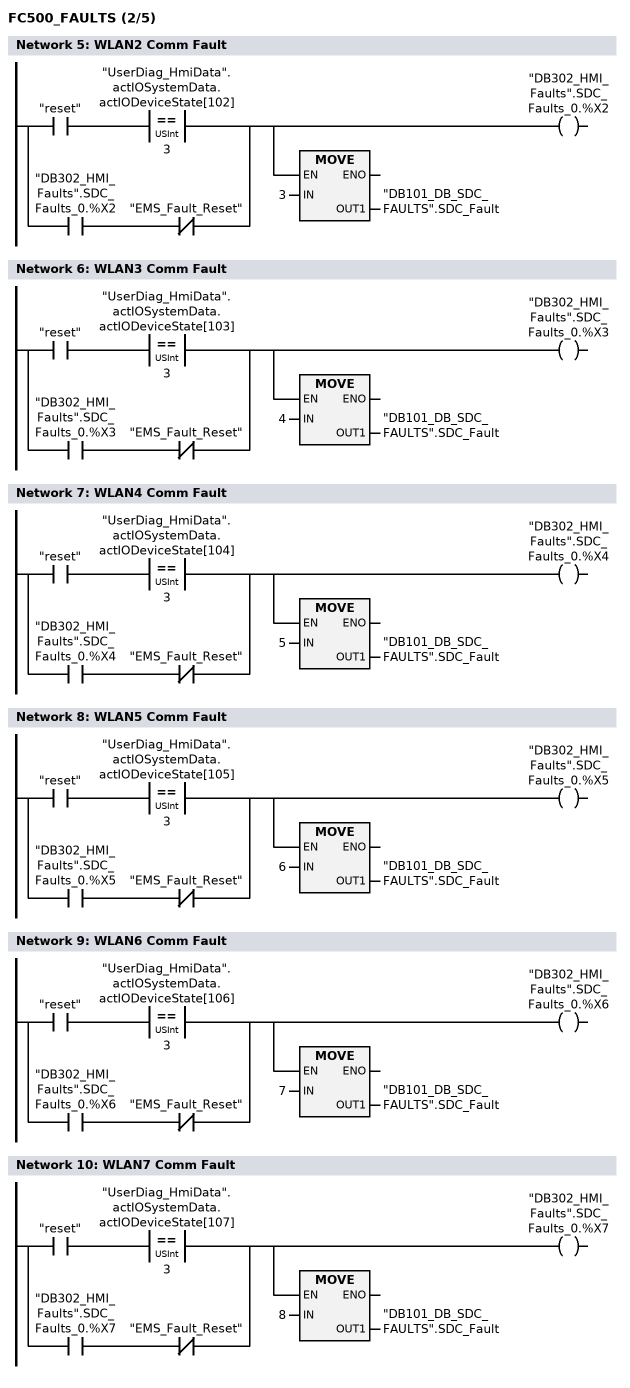
   RUNG wire#powerrail
      Contact( "reset" )
      { S7_Templates := "SrcType := USInt" } EQ_Contact(in1 := "UserDiag_HmiData".actIOSystemData.actIODeviceState[102], in2 := 3)
      wire#w1
      Coil( "DB302_HMI_Faults".SDC_Faults_0.%X2 )
   END_RUNG
   RUNG wire#powerrail
      Contact( "DB302_HMI_Faults".SDC_Faults_0.%X2 )
      I_Contact( "EMS_Fault_Reset" )
   END_RUNG wire#w1
   RUNG wire#w1
      Move(in := 3, out1 => "DB101_DB_SDC_FAULTS".SDC_Fault)
   END_RUNG
   // the same network as SCL:
   "DB302_HMI_Faults".SDC_Faults_0.%X2 := ("reset" AND ("UserDiag_HmiData".actIOSystemData.actIODeviceState[102] = 3)) OR ("DB302_HMI_Faults".SDC_Faults_0.%X2 AND NOT "EMS_Fault_Reset");
   IF "DB302_HMI_Faults".SDC_Faults_0.%X2 THEN "DB101_DB_SDC_FAULTS".SDC_Fault := 3; END_IF;
END_REGION

REGION Network 6: WLAN3 Comm Fault
   RUNG wire#powerrail
      Contact( "reset" )
      { S7_Templates := "SrcType := USInt" } EQ_Contact(in1 := "UserDiag_HmiData".actIOSystemData.actIODeviceState[103], in2 := 3)
      wire#w1
      Coil( "DB302_HMI_Faults".SDC_Faults_0.%X3 )
   END_RUNG
   RUNG wire#powerrail
      Contact( "DB302_HMI_Faults".SDC_Faults_0.%X3 )
      I_Contact( "EMS_Fault_Reset" )
   END_RUNG wire#w1
   RUNG wire#w1
      Move(in := 4, out1 => "DB101_DB_SDC_FAULTS".SDC_Fault)
   END_RUNG
   // the same network as SCL:
   "DB302_HMI_Faults".SDC_Faults_0.%X3 := ("reset" AND ("UserDiag_HmiData".actIOSystemData.actIODeviceState[103] = 3)) OR ("DB302_HMI_Faults".SDC_Faults_0.%X3 AND NOT "EMS_Fault_Reset");
   IF "DB302_HMI_Faults".SDC_Faults_0.%X3 THEN "DB101_DB_SDC_FAULTS".SDC_Fault := 4; END_IF;
END_REGION

REGION Network 7: WLAN4 Comm Fault
   RUNG wire#powerrail
      Contact( "reset" )
      { S7_Templates := "SrcType := USInt" } EQ_Contact(in1 := "UserDiag_HmiData".actIOSystemData.actIODeviceState[104], in2 := 3)
      wire#w1
      Coil( "DB302_HMI_Faults".SDC_Faults_0.%X4 )
   END_RUNG
   RUNG wire#powerrail
      Contact( "DB302_HMI_Faults".SDC_Faults_0.%X4 )
      I_Contact( "EMS_Fault_Reset" )
   END_RUNG wire#w1
   RUNG wire#w1
      Move(in := 5, out1 => "DB101_DB_SDC_FAULTS".SDC_Fault)
   END_RUNG
   // the same network as SCL:
   "DB302_HMI_Faults".SDC_Faults_0.%X4 := ("reset" AND ("UserDiag_HmiData".actIOSystemData.actIODeviceState[104] = 3)) OR ("DB302_HMI_Faults".SDC_Faults_0.%X4 AND NOT "EMS_Fault_Reset");
   IF "DB302_HMI_Faults".SDC_Faults_0.%X4 THEN "DB101_DB_SDC_FAULTS".SDC_Fault := 5; END_IF;
END_REGION

REGION Network 8: WLAN5 Comm Fault
   RUNG wire#powerrail
      Contact( "reset" )
      { S7_Templates := "SrcType := USInt" } EQ_Contact(in1 := "UserDiag_HmiData".actIOSystemData.actIODeviceState[105], in2 := 3)
      wire#w1
      Coil( "DB302_HMI_Faults".SDC_Faults_0.%X5 )
   END_RUNG
   RUNG wire#powerrail
      Contact( "DB302_HMI_Faults".SDC_Faults_0.%X5 )
      I_Contact( "EMS_Fault_Reset" )
   END_RUNG wire#w1
   RUNG wire#w1
      Move(in := 6, out1 => "DB101_DB_SDC_FAULTS".SDC_Fault)
   END_RUNG
   // the same network as SCL:
   "DB302_HMI_Faults".SDC_Faults_0.%X5 := ("reset" AND ("UserDiag_HmiData".actIOSystemData.actIODeviceState[105] = 3)) OR ("DB302_HMI_Faults".SDC_Faults_0.%X5 AND NOT "EMS_Fault_Reset");
   IF "DB302_HMI_Faults".SDC_Faults_0.%X5 THEN "DB101_DB_SDC_FAULTS".SDC_Fault := 6; END_IF;
END_REGION

REGION Network 9: WLAN6 Comm Fault
   RUNG wire#powerrail
      Contact( "reset" )
      { S7_Templates := "SrcType := USInt" } EQ_Contact(in1 := "UserDiag_HmiData".actIOSystemData.actIODeviceState[106], in2 := 3)
      wire#w1
      Coil( "DB302_HMI_Faults".SDC_Faults_0.%X6 )
   END_RUNG
   RUNG wire#powerrail
      Contact( "DB302_HMI_Faults".SDC_Faults_0.%X6 )
      I_Contact( "EMS_Fault_Reset" )
   END_RUNG wire#w1
   RUNG wire#w1
      Move(in := 7, out1 => "DB101_DB_SDC_FAULTS".SDC_Fault)
   END_RUNG
   // the same network as SCL:
   "DB302_HMI_Faults".SDC_Faults_0.%X6 := ("reset" AND ("UserDiag_HmiData".actIOSystemData.actIODeviceState[106] = 3)) OR ("DB302_HMI_Faults".SDC_Faults_0.%X6 AND NOT "EMS_Fault_Reset");
   IF "DB302_HMI_Faults".SDC_Faults_0.%X6 THEN "DB101_DB_SDC_FAULTS".SDC_Fault := 7; END_IF;
END_REGION

REGION Network 10: WLAN7 Comm Fault
   RUNG wire#powerrail
      Contact( "reset" )
      { S7_Templates := "SrcType := USInt" } EQ_Contact(in1 := "UserDiag_HmiData".actIOSystemData.actIODeviceState[107], in2 := 3)
      wire#w1
      Coil( "DB302_HMI_Faults".SDC_Faults_0.%X7 )
   END_RUNG
   RUNG wire#powerrail
      Contact( "DB302_HMI_Faults".SDC_Faults_0.%X7 )
      I_Contact( "EMS_Fault_Reset" )
   END_RUNG wire#w1
   RUNG wire#w1
      Move(in := 8, out1 => "DB101_DB_SDC_FAULTS".SDC_Fault)
   END_RUNG
   // the same network as SCL:
   "DB302_HMI_Faults".SDC_Faults_0.%X7 := ("reset" AND ("UserDiag_HmiData".actIOSystemData.actIODeviceState[107] = 3)) OR ("DB302_HMI_Faults".SDC_Faults_0.%X7 AND NOT "EMS_Fault_Reset");
   IF "DB302_HMI_Faults".SDC_Faults_0.%X7 THEN "DB101_DB_SDC_FAULTS".SDC_Fault := 8; END_IF;
END_REGION

REGION Network 11: WLAN8 Comm Fault
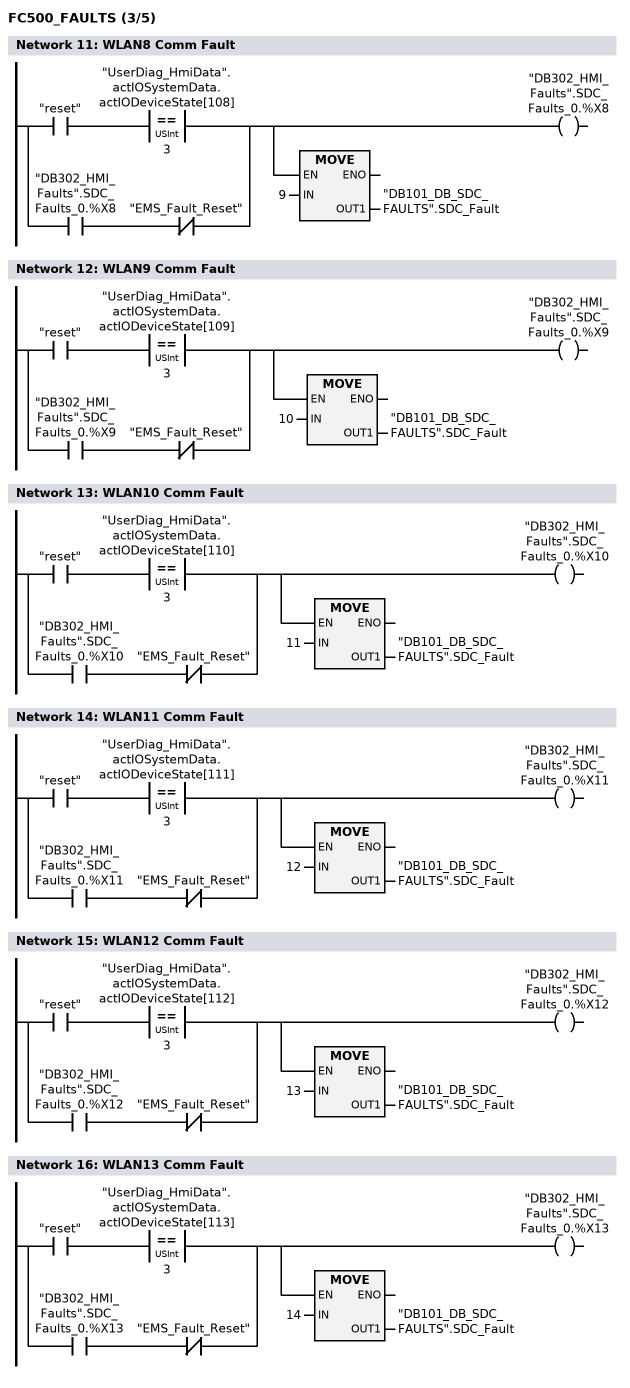
   RUNG wire#powerrail
      Contact( "reset" )
      { S7_Templates := "SrcType := USInt" } EQ_Contact(in1 := "UserDiag_HmiData".actIOSystemData.actIODeviceState[108], in2 := 3)
      wire#w1
      Coil( "DB302_HMI_Faults".SDC_Faults_0.%X8 )
   END_RUNG
   RUNG wire#powerrail
      Contact( "DB302_HMI_Faults".SDC_Faults_0.%X8 )
      I_Contact( "EMS_Fault_Reset" )
   END_RUNG wire#w1
   RUNG wire#w1
      Move(in := 9, out1 => "DB101_DB_SDC_FAULTS".SDC_Fault)
   END_RUNG
   // the same network as SCL:
   "DB302_HMI_Faults".SDC_Faults_0.%X8 := ("reset" AND ("UserDiag_HmiData".actIOSystemData.actIODeviceState[108] = 3)) OR ("DB302_HMI_Faults".SDC_Faults_0.%X8 AND NOT "EMS_Fault_Reset");
   IF "DB302_HMI_Faults".SDC_Faults_0.%X8 THEN "DB101_DB_SDC_FAULTS".SDC_Fault := 9; END_IF;
END_REGION

REGION Network 12: WLAN9 Comm Fault
   RUNG wire#powerrail
      Contact( "reset" )
      { S7_Templates := "SrcType := USInt" } EQ_Contact(in1 := "UserDiag_HmiData".actIOSystemData.actIODeviceState[109], in2 := 3)
      wire#w1
      Coil( "DB302_HMI_Faults".SDC_Faults_0.%X9 )
   END_RUNG
   RUNG wire#powerrail
      Contact( "DB302_HMI_Faults".SDC_Faults_0.%X9 )
      I_Contact( "EMS_Fault_Reset" )
   END_RUNG wire#w1
   RUNG wire#w1
      Move(in := 10, out1 => "DB101_DB_SDC_FAULTS".SDC_Fault)
   END_RUNG
   // the same network as SCL:
   "DB302_HMI_Faults".SDC_Faults_0.%X9 := ("reset" AND ("UserDiag_HmiData".actIOSystemData.actIODeviceState[109] = 3)) OR ("DB302_HMI_Faults".SDC_Faults_0.%X9 AND NOT "EMS_Fault_Reset");
   IF "DB302_HMI_Faults".SDC_Faults_0.%X9 THEN "DB101_DB_SDC_FAULTS".SDC_Fault := 10; END_IF;
END_REGION

REGION Network 13: WLAN10 Comm Fault
   RUNG wire#powerrail
      Contact( "reset" )
      { S7_Templates := "SrcType := USInt" } EQ_Contact(in1 := "UserDiag_HmiData".actIOSystemData.actIODeviceState[110], in2 := 3)
      wire#w1
      Coil( "DB302_HMI_Faults".SDC_Faults_0.%X10 )
   END_RUNG
   RUNG wire#powerrail
      Contact( "DB302_HMI_Faults".SDC_Faults_0.%X10 )
      I_Contact( "EMS_Fault_Reset" )
   END_RUNG wire#w1
   RUNG wire#w1
      Move(in := 11, out1 => "DB101_DB_SDC_FAULTS".SDC_Fault)
   END_RUNG
   // the same network as SCL:
   "DB302_HMI_Faults".SDC_Faults_0.%X10 := ("reset" AND ("UserDiag_HmiData".actIOSystemData.actIODeviceState[110] = 3)) OR ("DB302_HMI_Faults".SDC_Faults_0.%X10 AND NOT "EMS_Fault_Reset");
   IF "DB302_HMI_Faults".SDC_Faults_0.%X10 THEN "DB101_DB_SDC_FAULTS".SDC_Fault := 11; END_IF;
END_REGION

REGION Network 14: WLAN11 Comm Fault
   RUNG wire#powerrail
      Contact( "reset" )
      { S7_Templates := "SrcType := USInt" } EQ_Contact(in1 := "UserDiag_HmiData".actIOSystemData.actIODeviceState[111], in2 := 3)
      wire#w1
      Coil( "DB302_HMI_Faults".SDC_Faults_0.%X11 )
   END_RUNG
   RUNG wire#powerrail
      Contact( "DB302_HMI_Faults".SDC_Faults_0.%X11 )
      I_Contact( "EMS_Fault_Reset" )
   END_RUNG wire#w1
   RUNG wire#w1
      Move(in := 12, out1 => "DB101_DB_SDC_FAULTS".SDC_Fault)
   END_RUNG
   // the same network as SCL:
   "DB302_HMI_Faults".SDC_Faults_0.%X11 := ("reset" AND ("UserDiag_HmiData".actIOSystemData.actIODeviceState[111] = 3)) OR ("DB302_HMI_Faults".SDC_Faults_0.%X11 AND NOT "EMS_Fault_Reset");
   IF "DB302_HMI_Faults".SDC_Faults_0.%X11 THEN "DB101_DB_SDC_FAULTS".SDC_Fault := 12; END_IF;
END_REGION

REGION Network 15: WLAN12 Comm Fault
   RUNG wire#powerrail
      Contact( "reset" )
      { S7_Templates := "SrcType := USInt" } EQ_Contact(in1 := "UserDiag_HmiData".actIOSystemData.actIODeviceState[112], in2 := 3)
      wire#w1
      Coil( "DB302_HMI_Faults".SDC_Faults_0.%X12 )
   END_RUNG
   RUNG wire#powerrail
      Contact( "DB302_HMI_Faults".SDC_Faults_0.%X12 )
      I_Contact( "EMS_Fault_Reset" )
   END_RUNG wire#w1
   RUNG wire#w1
      Move(in := 13, out1 => "DB101_DB_SDC_FAULTS".SDC_Fault)
   END_RUNG
   // the same network as SCL:
   "DB302_HMI_Faults".SDC_Faults_0.%X12 := ("reset" AND ("UserDiag_HmiData".actIOSystemData.actIODeviceState[112] = 3)) OR ("DB302_HMI_Faults".SDC_Faults_0.%X12 AND NOT "EMS_Fault_Reset");
   IF "DB302_HMI_Faults".SDC_Faults_0.%X12 THEN "DB101_DB_SDC_FAULTS".SDC_Fault := 13; END_IF;
END_REGION

REGION Network 16: WLAN13 Comm Fault
   RUNG wire#powerrail
      Contact( "reset" )
      { S7_Templates := "SrcType := USInt" } EQ_Contact(in1 := "UserDiag_HmiData".actIOSystemData.actIODeviceState[113], in2 := 3)
      wire#w1
      Coil( "DB302_HMI_Faults".SDC_Faults_0.%X13 )
   END_RUNG
   RUNG wire#powerrail
      Contact( "DB302_HMI_Faults".SDC_Faults_0.%X13 )
      I_Contact( "EMS_Fault_Reset" )
   END_RUNG wire#w1
   RUNG wire#w1
      Move(in := 14, out1 => "DB101_DB_SDC_FAULTS".SDC_Fault)
   END_RUNG
   // the same network as SCL:
   "DB302_HMI_Faults".SDC_Faults_0.%X13 := ("reset" AND ("UserDiag_HmiData".actIOSystemData.actIODeviceState[113] = 3)) OR ("DB302_HMI_Faults".SDC_Faults_0.%X13 AND NOT "EMS_Fault_Reset");
   IF "DB302_HMI_Faults".SDC_Faults_0.%X13 THEN "DB101_DB_SDC_FAULTS".SDC_Fault := 14; END_IF;
END_REGION

REGION Network 17: WLAN14 Comm Fault
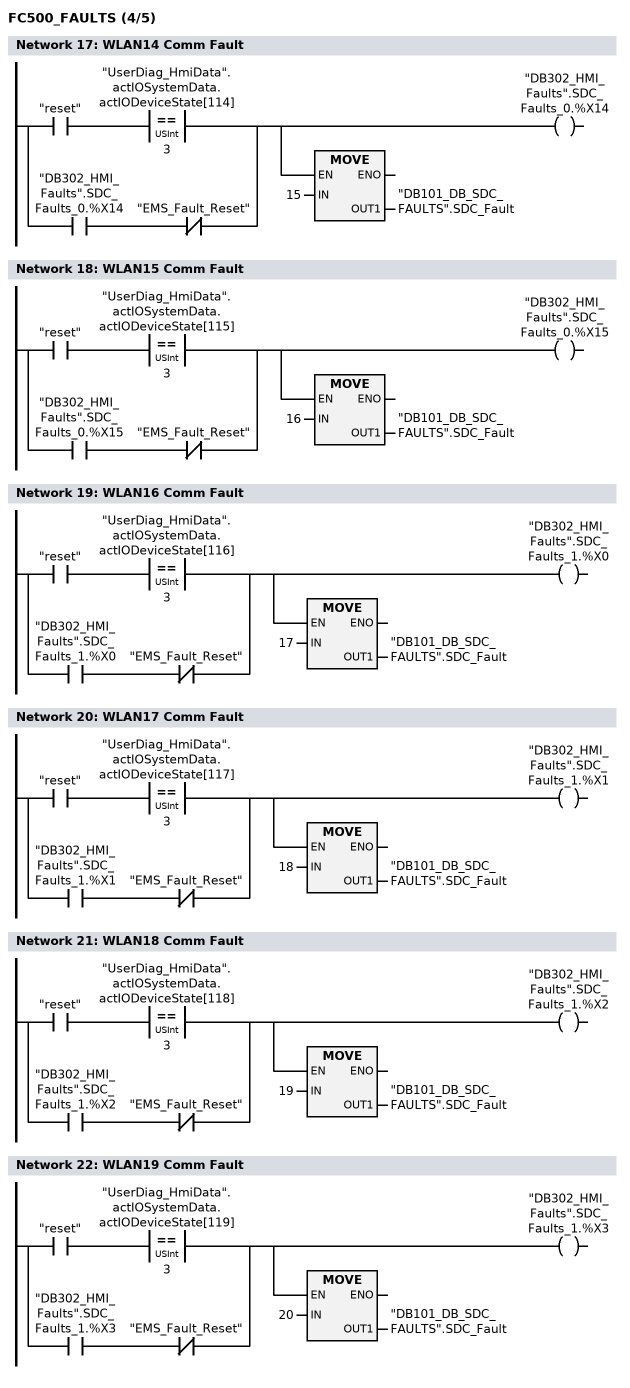
   RUNG wire#powerrail
      Contact( "reset" )
      { S7_Templates := "SrcType := USInt" } EQ_Contact(in1 := "UserDiag_HmiData".actIOSystemData.actIODeviceState[114], in2 := 3)
      wire#w1
      Coil( "DB302_HMI_Faults".SDC_Faults_0.%X14 )
   END_RUNG
   RUNG wire#powerrail
      Contact( "DB302_HMI_Faults".SDC_Faults_0.%X14 )
      I_Contact( "EMS_Fault_Reset" )
   END_RUNG wire#w1
   RUNG wire#w1
      Move(in := 15, out1 => "DB101_DB_SDC_FAULTS".SDC_Fault)
   END_RUNG
   // the same network as SCL:
   "DB302_HMI_Faults".SDC_Faults_0.%X14 := ("reset" AND ("UserDiag_HmiData".actIOSystemData.actIODeviceState[114] = 3)) OR ("DB302_HMI_Faults".SDC_Faults_0.%X14 AND NOT "EMS_Fault_Reset");
   IF "DB302_HMI_Faults".SDC_Faults_0.%X14 THEN "DB101_DB_SDC_FAULTS".SDC_Fault := 15; END_IF;
END_REGION

REGION Network 18: WLAN15 Comm Fault
   RUNG wire#powerrail
      Contact( "reset" )
      { S7_Templates := "SrcType := USInt" } EQ_Contact(in1 := "UserDiag_HmiData".actIOSystemData.actIODeviceState[115], in2 := 3)
      wire#w1
      Coil( "DB302_HMI_Faults".SDC_Faults_0.%X15 )
   END_RUNG
   RUNG wire#powerrail
      Contact( "DB302_HMI_Faults".SDC_Faults_0.%X15 )
      I_Contact( "EMS_Fault_Reset" )
   END_RUNG wire#w1
   RUNG wire#w1
      Move(in := 16, out1 => "DB101_DB_SDC_FAULTS".SDC_Fault)
   END_RUNG
   // the same network as SCL:
   "DB302_HMI_Faults".SDC_Faults_0.%X15 := ("reset" AND ("UserDiag_HmiData".actIOSystemData.actIODeviceState[115] = 3)) OR ("DB302_HMI_Faults".SDC_Faults_0.%X15 AND NOT "EMS_Fault_Reset");
   IF "DB302_HMI_Faults".SDC_Faults_0.%X15 THEN "DB101_DB_SDC_FAULTS".SDC_Fault := 16; END_IF;
END_REGION

REGION Network 19: WLAN16 Comm Fault
   RUNG wire#powerrail
      Contact( "reset" )
      { S7_Templates := "SrcType := USInt" } EQ_Contact(in1 := "UserDiag_HmiData".actIOSystemData.actIODeviceState[116], in2 := 3)
      wire#w1
      Coil( "DB302_HMI_Faults".SDC_Faults_1.%X0 )
   END_RUNG
   RUNG wire#powerrail
      Contact( "DB302_HMI_Faults".SDC_Faults_1.%X0 )
      I_Contact( "EMS_Fault_Reset" )
   END_RUNG wire#w1
   RUNG wire#w1
      Move(in := 17, out1 => "DB101_DB_SDC_FAULTS".SDC_Fault)
   END_RUNG
   // the same network as SCL:
   "DB302_HMI_Faults".SDC_Faults_1.%X0 := ("reset" AND ("UserDiag_HmiData".actIOSystemData.actIODeviceState[116] = 3)) OR ("DB302_HMI_Faults".SDC_Faults_1.%X0 AND NOT "EMS_Fault_Reset");
   IF "DB302_HMI_Faults".SDC_Faults_1.%X0 THEN "DB101_DB_SDC_FAULTS".SDC_Fault := 17; END_IF;
END_REGION

REGION Network 20: WLAN17 Comm Fault
   RUNG wire#powerrail
      Contact( "reset" )
      { S7_Templates := "SrcType := USInt" } EQ_Contact(in1 := "UserDiag_HmiData".actIOSystemData.actIODeviceState[117], in2 := 3)
      wire#w1
      Coil( "DB302_HMI_Faults".SDC_Faults_1.%X1 )
   END_RUNG
   RUNG wire#powerrail
      Contact( "DB302_HMI_Faults".SDC_Faults_1.%X1 )
      I_Contact( "EMS_Fault_Reset" )
   END_RUNG wire#w1
   RUNG wire#w1
      Move(in := 18, out1 => "DB101_DB_SDC_FAULTS".SDC_Fault)
   END_RUNG
   // the same network as SCL:
   "DB302_HMI_Faults".SDC_Faults_1.%X1 := ("reset" AND ("UserDiag_HmiData".actIOSystemData.actIODeviceState[117] = 3)) OR ("DB302_HMI_Faults".SDC_Faults_1.%X1 AND NOT "EMS_Fault_Reset");
   IF "DB302_HMI_Faults".SDC_Faults_1.%X1 THEN "DB101_DB_SDC_FAULTS".SDC_Fault := 18; END_IF;
END_REGION

REGION Network 21: WLAN18 Comm Fault
   RUNG wire#powerrail
      Contact( "reset" )
      { S7_Templates := "SrcType := USInt" } EQ_Contact(in1 := "UserDiag_HmiData".actIOSystemData.actIODeviceState[118], in2 := 3)
      wire#w1
      Coil( "DB302_HMI_Faults".SDC_Faults_1.%X2 )
   END_RUNG
   RUNG wire#powerrail
      Contact( "DB302_HMI_Faults".SDC_Faults_1.%X2 )
      I_Contact( "EMS_Fault_Reset" )
   END_RUNG wire#w1
   RUNG wire#w1
      Move(in := 19, out1 => "DB101_DB_SDC_FAULTS".SDC_Fault)
   END_RUNG
   // the same network as SCL:
   "DB302_HMI_Faults".SDC_Faults_1.%X2 := ("reset" AND ("UserDiag_HmiData".actIOSystemData.actIODeviceState[118] = 3)) OR ("DB302_HMI_Faults".SDC_Faults_1.%X2 AND NOT "EMS_Fault_Reset");
   IF "DB302_HMI_Faults".SDC_Faults_1.%X2 THEN "DB101_DB_SDC_FAULTS".SDC_Fault := 19; END_IF;
END_REGION

REGION Network 22: WLAN19 Comm Fault
   RUNG wire#powerrail
      Contact( "reset" )
      { S7_Templates := "SrcType := USInt" } EQ_Contact(in1 := "UserDiag_HmiData".actIOSystemData.actIODeviceState[119], in2 := 3)
      wire#w1
      Coil( "DB302_HMI_Faults".SDC_Faults_1.%X3 )
   END_RUNG
   RUNG wire#powerrail
      Contact( "DB302_HMI_Faults".SDC_Faults_1.%X3 )
      I_Contact( "EMS_Fault_Reset" )
   END_RUNG wire#w1
   RUNG wire#w1
      Move(in := 20, out1 => "DB101_DB_SDC_FAULTS".SDC_Fault)
   END_RUNG
   // the same network as SCL:
   "DB302_HMI_Faults".SDC_Faults_1.%X3 := ("reset" AND ("UserDiag_HmiData".actIOSystemData.actIODeviceState[119] = 3)) OR ("DB302_HMI_Faults".SDC_Faults_1.%X3 AND NOT "EMS_Fault_Reset");
   IF "DB302_HMI_Faults".SDC_Faults_1.%X3 THEN "DB101_DB_SDC_FAULTS".SDC_Fault := 20; END_IF;
END_REGION

REGION Network 23: Duplicate Carrier Fault
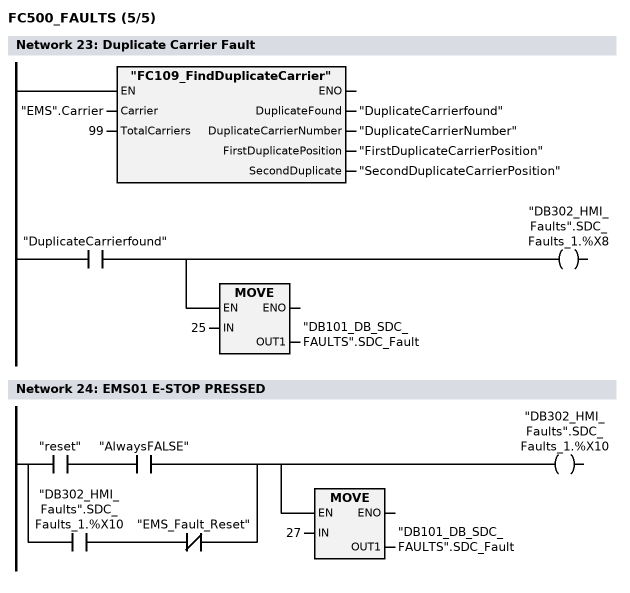
   RUNG wire#powerrail
      "FC109_FindDuplicateCarrier"(Carrier := "EMS".Carrier, TotalCarriers := 99, DuplicateFound => "DuplicateCarrierfound", DuplicateCarrierNumber => "DuplicateCarrierNumber", FirstDuplicatePosition => "FirstDuplicateCarrierPosition", SecondDuplicate => "SecondDuplicateCarrierPosition")
   END_RUNG
   RUNG wire#powerrail
      Contact( "DuplicateCarrierfound" )
      wire#w1
      Coil( "DB302_HMI_Faults".SDC_Faults_1.%X8 )
   END_RUNG
   RUNG wire#w1
      Move(in := 25, out1 => "DB101_DB_SDC_FAULTS".SDC_Fault)
   END_RUNG
   // the same network as SCL:
   "FC109_FindDuplicateCarrier"(Carrier := "EMS".Carrier,
                           TotalCarriers := 99,
                           DuplicateFound => "DuplicateCarrierfound",
                           DuplicateCarrierNumber => "DuplicateCarrierNumber",
                           FirstDuplicatePosition => "FirstDuplicateCarrierPosition",
                           SecondDuplicate => "SecondDuplicateCarrierPosition");
   "DB302_HMI_Faults".SDC_Faults_1.%X8 := "DuplicateCarrierfound";
   IF "DuplicateCarrierfound" THEN "DB101_DB_SDC_FAULTS".SDC_Fault := 25; END_IF;
END_REGION

REGION Network 24: EMS01 E-STOP PRESSED
   RUNG wire#powerrail
      Contact( "reset" )
      Contact( "AlwaysFALSE" )
      wire#w1
      Coil( "DB302_HMI_Faults".SDC_Faults_1.%X10 )
   END_RUNG
   RUNG wire#powerrail
      Contact( "DB302_HMI_Faults".SDC_Faults_1.%X10 )
      I_Contact( "EMS_Fault_Reset" )
   END_RUNG wire#w1
   RUNG wire#w1
      Move(in := 27, out1 => "DB101_DB_SDC_FAULTS".SDC_Fault)
   END_RUNG
   // the same network as SCL:
   "DB302_HMI_Faults".SDC_Faults_1.%X10 := ("reset" AND "AlwaysFALSE") OR ("DB302_HMI_Faults".SDC_Faults_1.%X10 AND NOT "EMS_Fault_Reset");
   IF "DB302_HMI_Faults".SDC_Faults_1.%X10 THEN "DB101_DB_SDC_FAULTS".SDC_Fault := 27; END_IF;
END_REGION
END_FUNCTION

FUNCTION "FC501_FAULTS  C1-C10" : Void   // FC501, LAD
{ S7_Optimized_Access := 'TRUE' }
VERSION : 0.1
BEGIN

REGION Network 1: CARRIER 1 FAULTS
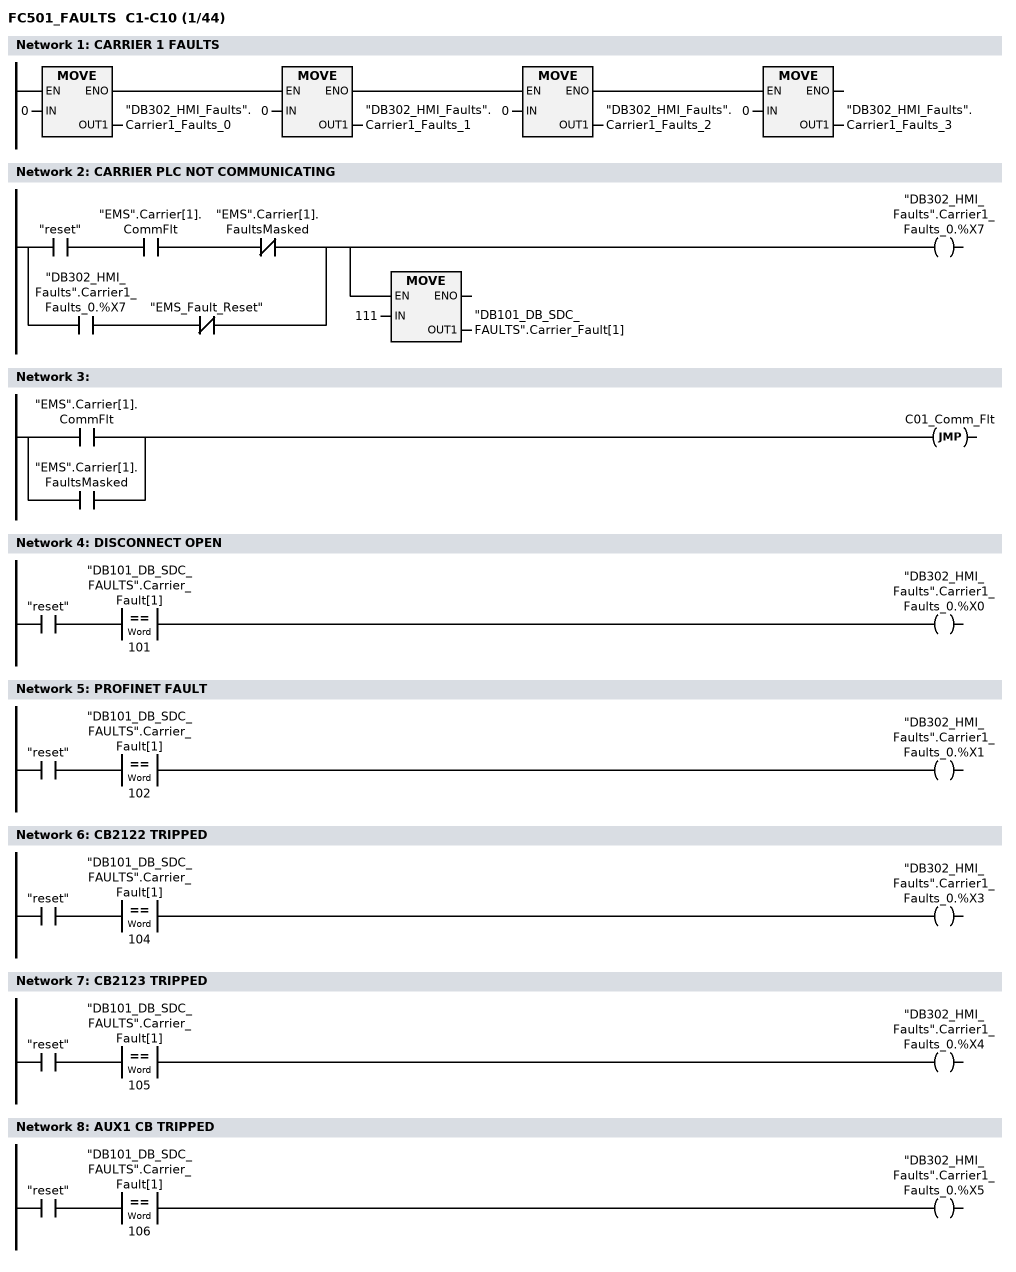
   RUNG wire#powerrail
      Move(in := 0, out1 => "DB302_HMI_Faults".Carrier1_Faults_0)
      Move(in := 0, out1 => "DB302_HMI_Faults".Carrier1_Faults_1)
      Move(in := 0, out1 => "DB302_HMI_Faults".Carrier1_Faults_2)
      Move(in := 0, out1 => "DB302_HMI_Faults".Carrier1_Faults_3)
   END_RUNG
   // the same network as SCL:
   "DB302_HMI_Faults".Carrier1_Faults_0 := 0;
   "DB302_HMI_Faults".Carrier1_Faults_1 := 0;
   "DB302_HMI_Faults".Carrier1_Faults_2 := 0;
   "DB302_HMI_Faults".Carrier1_Faults_3 := 0;
END_REGION

REGION Network 2: CARRIER PLC NOT COMMUNICATING
   RUNG wire#powerrail
      Contact( "reset" )
      Contact( "EMS".Carrier[1].CommFlt )
      I_Contact( "EMS".Carrier[1].FaultsMasked )
      wire#w1
      Coil( "DB302_HMI_Faults".Carrier1_Faults_0.%X7 )
   END_RUNG
   RUNG wire#powerrail
      Contact( "DB302_HMI_Faults".Carrier1_Faults_0.%X7 )
      I_Contact( "EMS_Fault_Reset" )
   END_RUNG wire#w1
   RUNG wire#w1
      Move(in := 111, out1 => "DB101_DB_SDC_FAULTS".Carrier_Fault[1])
   END_RUNG
   // the same network as SCL:
   "DB302_HMI_Faults".Carrier1_Faults_0.%X7 := ("reset" AND "EMS".Carrier[1].CommFlt AND NOT "EMS".Carrier[1].FaultsMasked) OR ("DB302_HMI_Faults".Carrier1_Faults_0.%X7 AND NOT "EMS_Fault_Reset");
   IF "DB302_HMI_Faults".Carrier1_Faults_0.%X7 THEN "DB101_DB_SDC_FAULTS".Carrier_Fault[1] := 111; END_IF;
END_REGION

REGION Network 3
   RUNG wire#powerrail
      Contact( "EMS".Carrier[1].CommFlt )
      wire#w1
      JumpCoil( C01_Comm_Flt )
   END_RUNG
   RUNG wire#powerrail
      Contact( "EMS".Carrier[1].FaultsMasked )
   END_RUNG wire#w1
   // the same network as SCL:
   IF "EMS".Carrier[1].CommFlt OR "EMS".Carrier[1].FaultsMasked THEN GOTO C01_Comm_Flt; END_IF;
END_REGION

REGION Network 4: DISCONNECT OPEN
   RUNG wire#powerrail
      Contact( "reset" )
      { S7_Templates := "SrcType := Word" } EQ_Contact(in1 := "DB101_DB_SDC_FAULTS".Carrier_Fault[1], in2 := 101)
      Coil( "DB302_HMI_Faults".Carrier1_Faults_0.%X0 )
   END_RUNG
   // the same network as SCL:
   "DB302_HMI_Faults".Carrier1_Faults_0.%X0 := "reset" AND ("DB101_DB_SDC_FAULTS".Carrier_Fault[1] = 101);
END_REGION

REGION Network 5: PROFINET FAULT
   RUNG wire#powerrail
      Contact( "reset" )
      { S7_Templates := "SrcType := Word" } EQ_Contact(in1 := "DB101_DB_SDC_FAULTS".Carrier_Fault[1], in2 := 102)
      Coil( "DB302_HMI_Faults".Carrier1_Faults_0.%X1 )
   END_RUNG
   // the same network as SCL:
   "DB302_HMI_Faults".Carrier1_Faults_0.%X1 := "reset" AND ("DB101_DB_SDC_FAULTS".Carrier_Fault[1] = 102);
END_REGION

REGION Network 6: CB2122 TRIPPED
   RUNG wire#powerrail
      Contact( "reset" )
      { S7_Templates := "SrcType := Word" } EQ_Contact(in1 := "DB101_DB_SDC_FAULTS".Carrier_Fault[1], in2 := 104)
      Coil( "DB302_HMI_Faults".Carrier1_Faults_0.%X3 )
   END_RUNG
   // the same network as SCL:
   "DB302_HMI_Faults".Carrier1_Faults_0.%X3 := "reset" AND ("DB101_DB_SDC_FAULTS".Carrier_Fault[1] = 104);
END_REGION

REGION Network 7: CB2123 TRIPPED
   RUNG wire#powerrail
      Contact( "reset" )
      { S7_Templates := "SrcType := Word" } EQ_Contact(in1 := "DB101_DB_SDC_FAULTS".Carrier_Fault[1], in2 := 105)
      Coil( "DB302_HMI_Faults".Carrier1_Faults_0.%X4 )
   END_RUNG
   // the same network as SCL:
   "DB302_HMI_Faults".Carrier1_Faults_0.%X4 := "reset" AND ("DB101_DB_SDC_FAULTS".Carrier_Fault[1] = 105);
END_REGION

REGION Network 8: AUX1 CB TRIPPED
   RUNG wire#powerrail
      Contact( "reset" )
      { S7_Templates := "SrcType := Word" } EQ_Contact(in1 := "DB101_DB_SDC_FAULTS".Carrier_Fault[1], in2 := 106)
      Coil( "DB302_HMI_Faults".Carrier1_Faults_0.%X5 )
   END_RUNG
   // the same network as SCL:
   "DB302_HMI_Faults".Carrier1_Faults_0.%X5 := "reset" AND ("DB101_DB_SDC_FAULTS".Carrier_Fault[1] = 106);
END_REGION

REGION Network 9: AUX2 CB TRIPPED
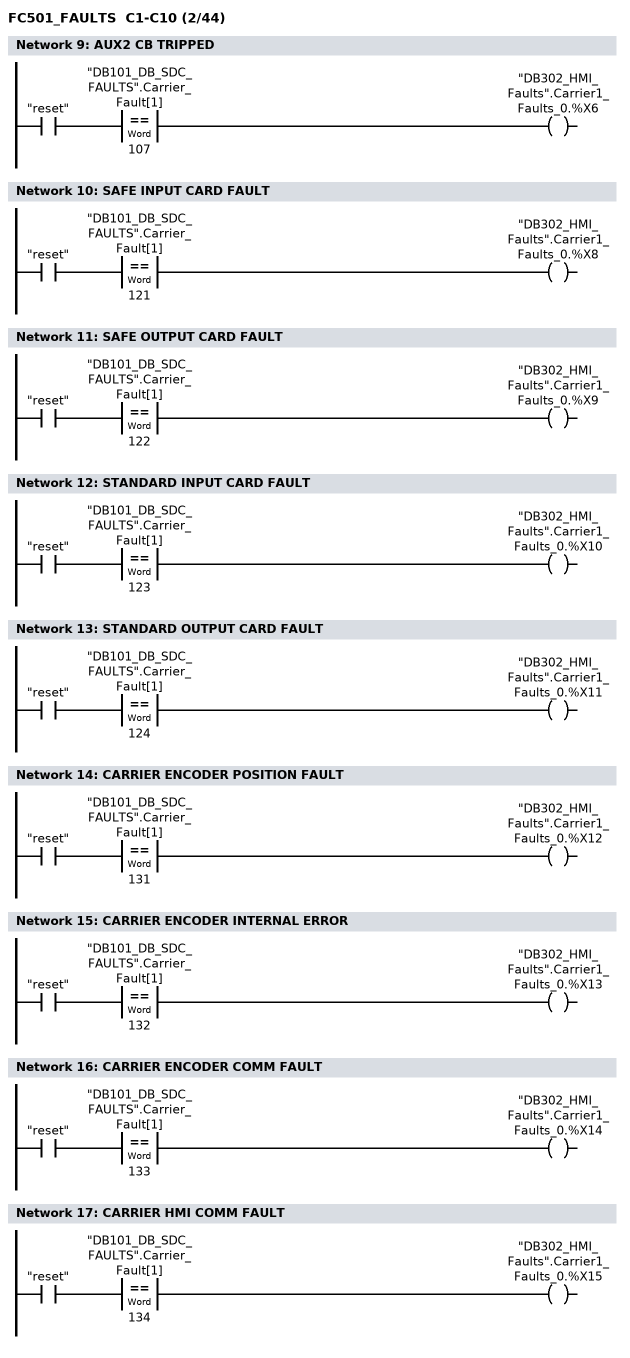
   RUNG wire#powerrail
      Contact( "reset" )
      { S7_Templates := "SrcType := Word" } EQ_Contact(in1 := "DB101_DB_SDC_FAULTS".Carrier_Fault[1], in2 := 107)
      Coil( "DB302_HMI_Faults".Carrier1_Faults_0.%X6 )
   END_RUNG
   // the same network as SCL:
   "DB302_HMI_Faults".Carrier1_Faults_0.%X6 := "reset" AND ("DB101_DB_SDC_FAULTS".Carrier_Fault[1] = 107);
END_REGION

REGION Network 10: SAFE INPUT CARD FAULT
   RUNG wire#powerrail
      Contact( "reset" )
      { S7_Templates := "SrcType := Word" } EQ_Contact(in1 := "DB101_DB_SDC_FAULTS".Carrier_Fault[1], in2 := 121)
      Coil( "DB302_HMI_Faults".Carrier1_Faults_0.%X8 )
   END_RUNG
   // the same network as SCL:
   "DB302_HMI_Faults".Carrier1_Faults_0.%X8 := "reset" AND ("DB101_DB_SDC_FAULTS".Carrier_Fault[1] = 121);
END_REGION

REGION Network 11: SAFE OUTPUT CARD FAULT
   RUNG wire#powerrail
      Contact( "reset" )
      { S7_Templates := "SrcType := Word" } EQ_Contact(in1 := "DB101_DB_SDC_FAULTS".Carrier_Fault[1], in2 := 122)
      Coil( "DB302_HMI_Faults".Carrier1_Faults_0.%X9 )
   END_RUNG
   // the same network as SCL:
   "DB302_HMI_Faults".Carrier1_Faults_0.%X9 := "reset" AND ("DB101_DB_SDC_FAULTS".Carrier_Fault[1] = 122);
END_REGION

REGION Network 12: STANDARD INPUT CARD FAULT
   RUNG wire#powerrail
      Contact( "reset" )
      { S7_Templates := "SrcType := Word" } EQ_Contact(in1 := "DB101_DB_SDC_FAULTS".Carrier_Fault[1], in2 := 123)
      Coil( "DB302_HMI_Faults".Carrier1_Faults_0.%X10 )
   END_RUNG
   // the same network as SCL:
   "DB302_HMI_Faults".Carrier1_Faults_0.%X10 := "reset" AND ("DB101_DB_SDC_FAULTS".Carrier_Fault[1] = 123);
END_REGION

REGION Network 13: STANDARD OUTPUT CARD FAULT
   RUNG wire#powerrail
      Contact( "reset" )
      { S7_Templates := "SrcType := Word" } EQ_Contact(in1 := "DB101_DB_SDC_FAULTS".Carrier_Fault[1], in2 := 124)
      Coil( "DB302_HMI_Faults".Carrier1_Faults_0.%X11 )
   END_RUNG
   // the same network as SCL:
   "DB302_HMI_Faults".Carrier1_Faults_0.%X11 := "reset" AND ("DB101_DB_SDC_FAULTS".Carrier_Fault[1] = 124);
END_REGION

REGION Network 14: CARRIER ENCODER POSITION FAULT
   RUNG wire#powerrail
      Contact( "reset" )
      { S7_Templates := "SrcType := Word" } EQ_Contact(in1 := "DB101_DB_SDC_FAULTS".Carrier_Fault[1], in2 := 131)
      Coil( "DB302_HMI_Faults".Carrier1_Faults_0.%X12 )
   END_RUNG
   // the same network as SCL:
   "DB302_HMI_Faults".Carrier1_Faults_0.%X12 := "reset" AND ("DB101_DB_SDC_FAULTS".Carrier_Fault[1] = 131);
END_REGION

REGION Network 15: CARRIER ENCODER INTERNAL ERROR
   RUNG wire#powerrail
      Contact( "reset" )
      { S7_Templates := "SrcType := Word" } EQ_Contact(in1 := "DB101_DB_SDC_FAULTS".Carrier_Fault[1], in2 := 132)
      Coil( "DB302_HMI_Faults".Carrier1_Faults_0.%X13 )
   END_RUNG
   // the same network as SCL:
   "DB302_HMI_Faults".Carrier1_Faults_0.%X13 := "reset" AND ("DB101_DB_SDC_FAULTS".Carrier_Fault[1] = 132);
END_REGION

REGION Network 16: CARRIER ENCODER COMM FAULT
   RUNG wire#powerrail
      Contact( "reset" )
      { S7_Templates := "SrcType := Word" } EQ_Contact(in1 := "DB101_DB_SDC_FAULTS".Carrier_Fault[1], in2 := 133)
      Coil( "DB302_HMI_Faults".Carrier1_Faults_0.%X14 )
   END_RUNG
   // the same network as SCL:
   "DB302_HMI_Faults".Carrier1_Faults_0.%X14 := "reset" AND ("DB101_DB_SDC_FAULTS".Carrier_Fault[1] = 133);
END_REGION

REGION Network 17: CARRIER HMI COMM FAULT
   RUNG wire#powerrail
      Contact( "reset" )
      { S7_Templates := "SrcType := Word" } EQ_Contact(in1 := "DB101_DB_SDC_FAULTS".Carrier_Fault[1], in2 := 134)
      Coil( "DB302_HMI_Faults".Carrier1_Faults_0.%X15 )
   END_RUNG
   // the same network as SCL:
   "DB302_HMI_Faults".Carrier1_Faults_0.%X15 := "reset" AND ("DB101_DB_SDC_FAULTS".Carrier_Fault[1] = 134);
END_REGION

REGION Network 18: CARRIER CRASH DETECTION FAULT